// TIA Portal project "FS-DS-09" (V16) (continued)
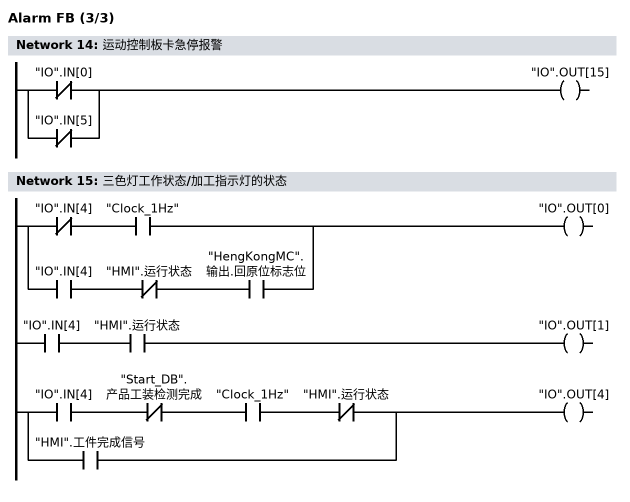
   RUNG wire#powerrail
      I_Contact( "IO".IN[0] )
      wire#w1
      Coil( "IO".OUT[15] )
   END_RUNG
   RUNG wire#powerrail
      I_Contact( "IO".IN[5] )
   END_RUNG wire#w1
   // the same network as SCL:
   "IO".OUT[15] := NOT "IO".IN[0] OR NOT "IO".IN[5];
END_REGION

REGION Network 15: 三色灯工作状态/加工指示灯的状态
   RUNG wire#powerrail
      I_Contact( "IO".IN[4] )
      Contact( "Clock_1Hz" )
      wire#w1
      Coil( "IO".OUT[0] )
   END_RUNG
   RUNG wire#powerrail
      Contact( "IO".IN[4] )
      I_Contact( "HMI".运行状态 )
      Contact( "HengKongMC".输出.回原位标志位 )
   END_RUNG wire#w1
   RUNG wire#powerrail
      Contact( "IO".IN[4] )
      Contact( "HMI".运行状态 )
      Coil( "IO".OUT[1] )
   END_RUNG
   RUNG wire#powerrail
      Contact( "IO".IN[4] )
      I_Contact( "Start_DB".产品工装检测完成 )
      Contact( "Clock_1Hz" )
      I_Contact( "HMI".运行状态 )
      wire#w2
      Coil( "IO".OUT[4] )
   END_RUNG
   RUNG wire#powerrail
      Contact( "HMI".工件完成信号 )
   END_RUNG wire#w2
   // the same network as SCL:
   "IO".OUT[0] := (NOT "IO".IN[4] AND "Clock_1Hz") OR ("IO".IN[4] AND NOT "HMI".运行状态 AND "HengKongMC".输出.回原位标志位);
   "IO".OUT[1] := "IO".IN[4] AND "HMI".运行状态;
   "IO".OUT[4] := ("IO".IN[4] AND NOT "Start_DB".产品工装检测完成 AND "Clock_1Hz" AND NOT "HMI".运行状态) OR "HMI".工件完成信号;
END_REGION
END_FUNCTION_BLOCK

// folder: Control

FUNCTION_BLOCK "Control FB"   // FB2, LAD
{ S7_Optimized_Access := 'TRUE' }
VERSION : 0.1
   VAR
      功能块_Instance : "AM/UM";
      功能块_Instance_1 : "AM/UM";
      功能块_Instance_2 : "AM/UM";
      功能块_Instance_3 : "AM/UM";
      功能块_Instance_4 : "AM/UM";
      功能块_Instance_5 : "AM/UM";
      功能块_Instance_6 : "AM/UM";
      功能块_Instance_7 : "AM/UM";
      IEC_Timer_0_Instance : TON_TIME;
      F_TRIG_Instance : F_TRIG;
      "AM/UM_1_Instance" : "AM/UM_1";
   END_VAR
BEGIN

REGION Network 1: Y1供料器有料输出
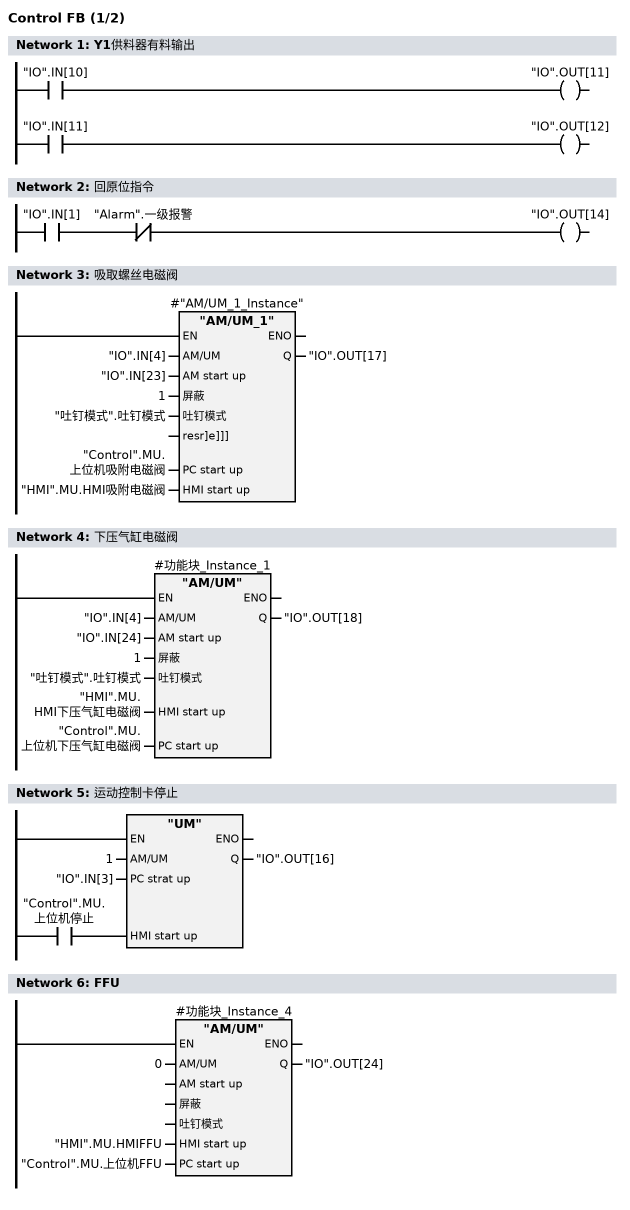
   RUNG wire#powerrail
      Contact( "IO".IN[10] )
      Coil( "IO".OUT[11] )
   END_RUNG
   RUNG wire#powerrail
      Contact( "IO".IN[11] )
      Coil( "IO".OUT[12] )
   END_RUNG
   // the same network as SCL:
   "IO".OUT[11] := "IO".IN[10];
   "IO".OUT[12] := "IO".IN[11];
END_REGION

REGION Network 2: 回原位指令
   RUNG wire#powerrail
      Contact( "IO".IN[1] )
      I_Contact( "Alarm".一级报警 )
      Coil( "IO".OUT[14] )
   END_RUNG
   // the same network as SCL:
   "IO".OUT[14] := "IO".IN[1] AND NOT "Alarm".一级报警;
END_REGION

REGION Network 3: 吸取螺丝电磁阀
   RUNG wire#powerrail
      #"AM/UM_1_Instance"("AM/UM" := "IO".IN[4], "AM start up" := "IO".IN[23], 屏蔽 := 1, 吐钉模式 := "吐钉模式".吐钉模式, "PC start up" := "Control".MU.上位机吸附电磁阀, "HMI start up" := "HMI".MU.HMI吸附电磁阀, Q => "IO".OUT[17], "resr]e]]]" :=)
   END_RUNG
   // the same network as SCL:
   #"AM/UM_1_Instance"("AM/UM" := "IO".IN[4],   // "AM/UM_1"
                       "AM start up" := "IO".IN[23],
                       屏蔽 := 1,
                       吐钉模式 := "吐钉模式".吐钉模式,
                       "PC start up" := "Control".MU.上位机吸附电磁阀,
                       "HMI start up" := "HMI".MU.HMI吸附电磁阀,
                       Q => "IO".OUT[17]);
END_REGION

REGION Network 4: 下压气缸电磁阀
   RUNG wire#powerrail
      #功能块_Instance_1("AM/UM" := "IO".IN[4], "AM start up" := "IO".IN[24], 屏蔽 := 1, 吐钉模式 := "吐钉模式".吐钉模式, "HMI start up" := "HMI".MU.HMI下压气缸电磁阀, "PC start up" := "Control".MU.上位机下压气缸电磁阀, Q => "IO".OUT[18])
   END_RUNG
   // the same network as SCL:
   #功能块_Instance_1("AM/UM" := "IO".IN[4],   // "AM/UM"
                   "AM start up" := "IO".IN[24],
                   屏蔽 := 1,
                   吐钉模式 := "吐钉模式".吐钉模式,
                   "HMI start up" := "HMI".MU.HMI下压气缸电磁阀,
                   "PC start up" := "Control".MU.上位机下压气缸电磁阀,
                   Q => "IO".OUT[18]);
END_REGION

REGION Network 5: 运动控制卡停止
   RUNG wire#powerrail
      "UM"("HMI start up" := wire#w1, "AM/UM" := 1, "PC strat up" := "IO".IN[3], Q => "IO".OUT[16])
   END_RUNG
   RUNG wire#powerrail
      Contact( "Control".MU.上位机停止 )
   END_RUNG wire#w1
   // the same network as SCL:
   "UM"("AM/UM" := 1, "PC strat up" := "IO".IN[3], "HMI start up" := "Control".MU.上位机停止, Q => "IO".OUT[16]);
END_REGION

REGION Network 6: FFU
   RUNG wire#powerrail
      #功能块_Instance_4("AM/UM" := 0, "AM start up" :=, 屏蔽 :=, 吐钉模式 :=, "HMI start up" := "HMI".MU.HMIFFU, "PC start up" := "Control".MU.上位机FFU, Q => "IO".OUT[24])
   END_RUNG
   // the same network as SCL:
   #功能块_Instance_4("AM/UM" := 0,   // "AM/UM"
                   "HMI start up" := "HMI".MU.HMIFFU,
                   "PC start up" := "Control".MU.上位机FFU,
                   Q => "IO".OUT[24]);
END_REGION

REGION Network 7: 照明
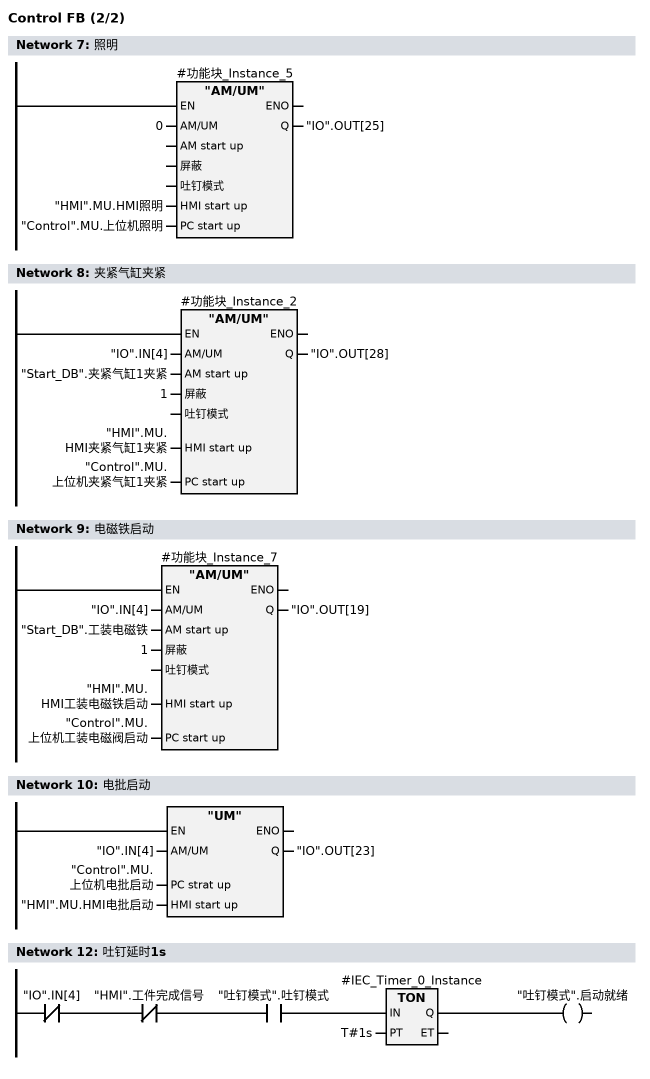
   RUNG wire#powerrail
      #功能块_Instance_5("AM/UM" := 0, "AM start up" :=, 屏蔽 :=, 吐钉模式 :=, "HMI start up" := "HMI".MU.HMI照明, "PC start up" := "Control".MU.上位机照明, Q => "IO".OUT[25])
   END_RUNG
   // the same network as SCL:
   #功能块_Instance_5("AM/UM" := 0,   // "AM/UM"
                   "HMI start up" := "HMI".MU.HMI照明,
                   "PC start up" := "Control".MU.上位机照明,
                   Q => "IO".OUT[25]);
END_REGION

REGION Network 8: 夹紧气缸夹紧
   RUNG wire#powerrail
      #功能块_Instance_2("AM/UM" := "IO".IN[4], "AM start up" := "Start_DB".夹紧气缸1夹紧, 屏蔽 := 1, 吐钉模式 :=, "HMI start up" := "HMI".MU.HMI夹紧气缸1夹紧, "PC start up" := "Control".MU.上位机夹紧气缸1夹紧, Q => "IO".OUT[28])
   END_RUNG
   // the same network as SCL:
   #功能块_Instance_2("AM/UM" := "IO".IN[4],   // "AM/UM"
                   "AM start up" := "Start_DB".夹紧气缸1夹紧,
                   屏蔽 := 1,
                   "HMI start up" := "HMI".MU.HMI夹紧气缸1夹紧,
                   "PC start up" := "Control".MU.上位机夹紧气缸1夹紧,
                   Q => "IO".OUT[28]);
END_REGION

REGION Network 9: 电磁铁启动
   RUNG wire#powerrail
      #功能块_Instance_7("AM/UM" := "IO".IN[4], "AM start up" := "Start_DB".工装电磁铁, 屏蔽 := 1, 吐钉模式 :=, "HMI start up" := "HMI".MU.HMI工装电磁铁启动, "PC start up" := "Control".MU.上位机工装电磁阀启动, Q => "IO".OUT[19])
   END_RUNG
   // the same network as SCL:
   #功能块_Instance_7("AM/UM" := "IO".IN[4],   // "AM/UM"
                   "AM start up" := "Start_DB".工装电磁铁,
                   屏蔽 := 1,
                   "HMI start up" := "HMI".MU.HMI工装电磁铁启动,
                   "PC start up" := "Control".MU.上位机工装电磁阀启动,
                   Q => "IO".OUT[19]);
END_REGION

REGION Network 10: 电批启动
   RUNG wire#powerrail
      "UM"("AM/UM" := "IO".IN[4], "PC strat up" := "Control".MU.上位机电批启动, "HMI start up" := "HMI".MU.HMI电批启动, Q => "IO".OUT[23])
   END_RUNG
   // the same network as SCL:
   "UM"("AM/UM" := "IO".IN[4],
        "PC strat up" := "Control".MU.上位机电批启动,
        "HMI start up" := "HMI".MU.HMI电批启动,
        Q => "IO".OUT[23]);
END_REGION

REGION Network 12: 吐钉延时1s
   #IEC_Timer_0_Instance(IN := NOT "IO".IN[4] AND NOT "HMI".工件完成信号 AND "吐钉模式".吐钉模式, PT := T#1s);   // TON
   "吐钉模式".启动就绪 := #IEC_Timer_0_Instance.Q;
END_REGION

REGION Network 13 (SCL): 完成后 复位
   #F_TRIG_Instance(CLK:="HengKongMC".输出.下压气缸信号,
                    Q=>"吐钉模式".下压气缸复位信号);
   IF "吐钉模式".下压气缸复位信号 OR  "IO".IN[1] THEN
       "吐钉模式".吐钉模式 := 0;
   END_IF;
END_REGION
END_FUNCTION_BLOCK

FUNCTION_BLOCK "Start"   // FB4, LAD
{ S7_Optimized_Access := 'TRUE' }
VERSION : 0.1
   VAR_OUTPUT
      夹紧气缸1夹紧 : Bool;
      夹紧气缸2夹紧 : Bool;
      工装电磁铁 : Bool;
   END_VAR
   VAR
      产品工装检测完成 : Bool;
      气缸夹紧完成 : Bool;
      P1 : Bool;
      P2 : Bool;
      RecipeExport_Instance : RecipeExport;
      RecipeImport_Instance : RecipeImport;
   END_VAR
   VAR_TEMP   // added for the SCL form of the ladder/FBD networks
      _w1 : Bool;
      _w2 : Bool;
   END_VAR
BEGIN

REGION Network 1: 启动1序/停止序
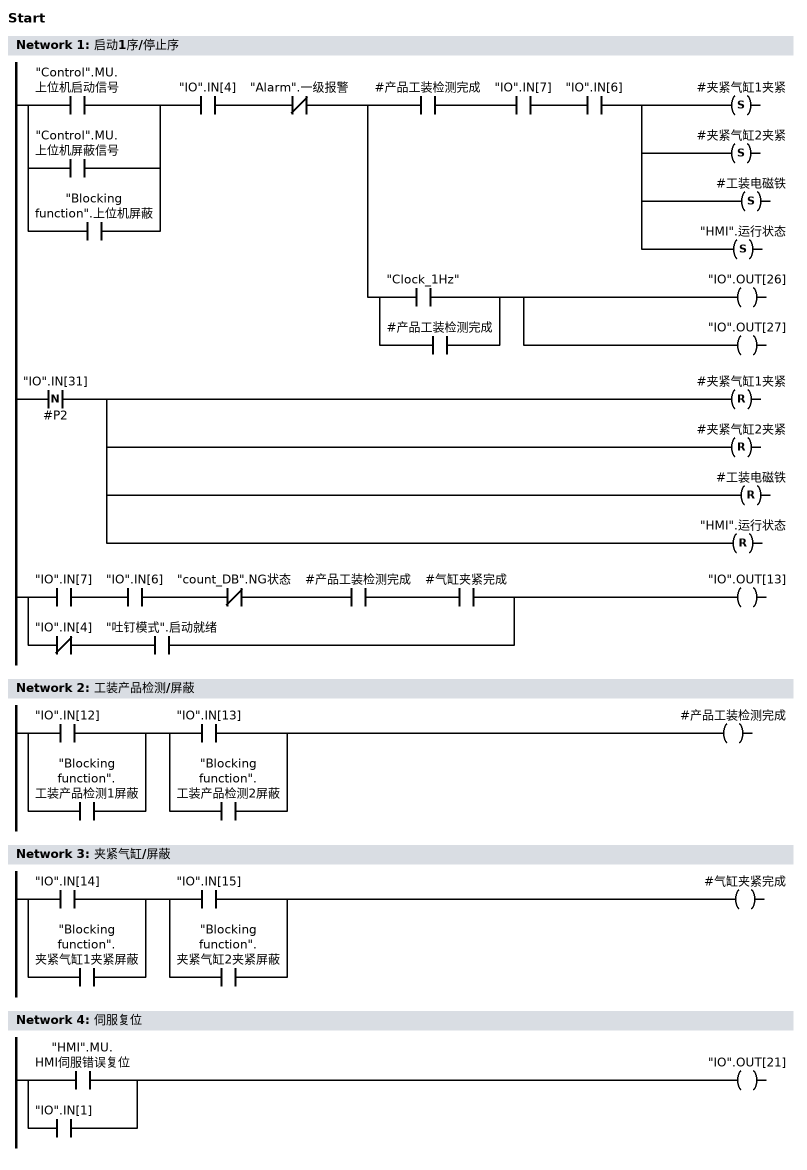
   RUNG wire#powerrail
      Contact( "Control".MU.上位机启动信号 )
      wire#w1
      Contact( "IO".IN[4] )
      I_Contact( "Alarm".一级报警 )
      wire#w2
      Contact( #产品工装检测完成 )
      Contact( "IO".IN[7] )
      Contact( "IO".IN[6] )
      wire#w3
      S_Coil( #夹紧气缸1夹紧 )
   END_RUNG
   RUNG wire#powerrail
      Contact( "Control".MU.上位机屏蔽信号 )
   END_RUNG wire#w1
   RUNG wire#powerrail
      Contact( "Blocking function".上位机屏蔽 )
   END_RUNG wire#w1
   RUNG wire#w3
      S_Coil( #夹紧气缸2夹紧 )
   END_RUNG
   RUNG wire#w3
      S_Coil( #工装电磁铁 )
   END_RUNG
   RUNG wire#w3
      S_Coil( "HMI".运行状态 )
   END_RUNG
   RUNG wire#w2
      Contact( "Clock_1Hz" )
      wire#w4
      Coil( "IO".OUT[26] )
   END_RUNG
   RUNG wire#w2
      Contact( #产品工装检测完成 )
   END_RUNG wire#w4
   RUNG wire#w4
      Coil( "IO".OUT[27] )
   END_RUNG
   RUNG wire#powerrail
      N_Contact(operand := "IO".IN[31], bit := #P2)
      wire#w5
      R_Coil( #夹紧气缸1夹紧 )
   END_RUNG
   RUNG wire#w5
      R_Coil( #夹紧气缸2夹紧 )
   END_RUNG
   RUNG wire#w5
      R_Coil( #工装电磁铁 )
   END_RUNG
   RUNG wire#w5
      R_Coil( "HMI".运行状态 )
   END_RUNG
   RUNG wire#powerrail
      Contact( "IO".IN[7] )
      Contact( "IO".IN[6] )
      I_Contact( "count_DB".NG状态 )
      Contact( #产品工装检测完成 )
      Contact( #气缸夹紧完成 )
      wire#w6
      Coil( "IO".OUT[13] )
   END_RUNG
   RUNG wire#powerrail
      I_Contact( "IO".IN[4] )
      Contact( "吐钉模式".启动就绪 )
   END_RUNG wire#w6
   // the same network as SCL:
   #_w1 := ("Control".MU.上位机启动信号 OR "Control".MU.上位机屏蔽信号 OR "Blocking function".上位机屏蔽) AND "IO".IN[4] AND NOT "Alarm".一级报警;
   IF #_w1 AND #产品工装检测完成 AND "IO".IN[7] AND "IO".IN[6] THEN
       #夹紧气缸1夹紧 := TRUE;
       #夹紧气缸2夹紧 := TRUE;
       #工装电磁铁 := TRUE;
       "HMI".运行状态 := TRUE;
   END_IF;
   "IO".OUT[26] := #_w1 AND ("Clock_1Hz" OR #产品工装检测完成);
   "IO".OUT[27] := #_w1 AND ("Clock_1Hz" OR #产品工装检测完成);
   #_w2 := NOT "IO".IN[31] AND #P2;   // falling edge of "IO".IN[31]
   #P2 := "IO".IN[31];
   IF #_w2 THEN
       #夹紧气缸1夹紧 := FALSE;
       #夹紧气缸2夹紧 := FALSE;
       #工装电磁铁 := FALSE;
       "HMI".运行状态 := FALSE;
   END_IF;
   "IO".OUT[13] := ("IO".IN[7] AND "IO".IN[6] AND NOT "count_DB".NG状态 AND #产品工装检测完成 AND #气缸夹紧完成) OR (NOT "IO".IN[4] AND "吐钉模式".启动就绪);
END_REGION

REGION Network 2: 工装产品检测/屏蔽
   RUNG wire#powerrail
      Contact( "IO".IN[12] )
      wire#w1
      Contact( "IO".IN[13] )
      wire#w2
      Coil( #产品工装检测完成 )
   END_RUNG
   RUNG wire#powerrail
      Contact( "Blocking function".工装产品检测1屏蔽 )
   END_RUNG wire#w1
   RUNG wire#w1
      Contact( "Blocking function".工装产品检测2屏蔽 )
   END_RUNG wire#w2
   // the same network as SCL:
   #产品工装检测完成 := ("IO".IN[12] OR "Blocking function".工装产品检测1屏蔽) AND ("IO".IN[13] OR "Blocking function".工装产品检测2屏蔽);
END_REGION

REGION Network 3: 夹紧气缸/屏蔽
   RUNG wire#powerrail
      Contact( "IO".IN[14] )
      wire#w1
      Contact( "IO".IN[15] )
      wire#w2
      Coil( #气缸夹紧完成 )
   END_RUNG
   RUNG wire#powerrail
      Contact( "Blocking function".夹紧气缸1夹紧屏蔽 )
   END_RUNG wire#w1
   RUNG wire#w1
      Contact( "Blocking function".夹紧气缸2夹紧屏蔽 )
   END_RUNG wire#w2
   // the same network as SCL:
   #气缸夹紧完成 := ("IO".IN[14] OR "Blocking function".夹紧气缸1夹紧屏蔽) AND ("IO".IN[15] OR "Blocking function".夹紧气缸2夹紧屏蔽);
END_REGION

REGION Network 4: 伺服复位
   RUNG wire#powerrail
      Contact( "HMI".MU.HMI伺服错误复位 )
      wire#w1
      Coil( "IO".OUT[21] )
   END_RUNG
   RUNG wire#powerrail
      Contact( "IO".IN[1] )
   END_RUNG wire#w1
   // the same network as SCL:
   "IO".OUT[21] := "HMI".MU.HMI伺服错误复位 OR "IO".IN[1];
END_REGION
END_FUNCTION_BLOCK

FUNCTION_BLOCK "AM/UM"   // FB5, LAD
{ S7_Optimized_Access := 'TRUE' }
VERSION : 0.1
   VAR_INPUT
      "AM/UM" : Bool;   // 手动自动
      "AM start up" : Bool;   // 自动启动
      屏蔽 : Bool;   // 屏蔽0
      吐钉模式 : Bool;
   END_VAR
   VAR_OUTPUT
      Q : Bool;   // 功能输出
   END_VAR
   VAR_IN_OUT
      "HMI start up" : Bool;   // HMI启动
      "PC start up" : Bool;   // 上位机启动
   END_VAR
   VAR
      F_TRIG_Instance : F_TRIG;
   END_VAR
BEGIN

REGION Network 1: 功能输出
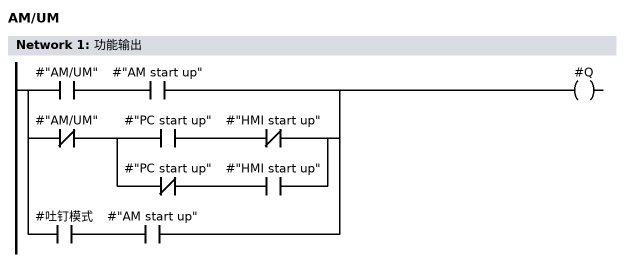
   RUNG wire#powerrail
      Contact( #"AM/UM" )
      Contact( #"AM start up" )
      wire#w1
      Coil( #Q )
   END_RUNG
   RUNG wire#powerrail
      I_Contact( #"AM/UM" )
      wire#w2
      Contact( #"PC start up" )
      I_Contact( #"HMI start up" )
   END_RUNG wire#w1
   RUNG wire#w2
      I_Contact( #"PC start up" )
      Contact( #"HMI start up" )
   END_RUNG wire#w1
   RUNG wire#powerrail
      Contact( #吐钉模式 )
      Contact( #"AM start up" )
   END_RUNG wire#w1
   // the same network as SCL:
   #Q := (#"AM/UM" AND #"AM start up") OR (NOT #"AM/UM" AND ((#"PC start up" AND NOT #"HMI start up") OR (NOT #"PC start up" AND #"HMI start up"))) OR (#吐钉模式 AND #"AM start up");
END_REGION

REGION Network 2 (SCL): HMI启动
   IF #屏蔽 THEN
       IF #"AM/UM" = 1 THEN
           #"HMI start up" := 0;
           #"PC start up":=0
           ;
       END_IF;
   END_IF;
END_REGION
END_FUNCTION_BLOCK

FUNCTION_BLOCK "count"   // FB7, LAD
{ S7_Optimized_Access := 'TRUE' }
VERSION : 0.1
// 计数OK/NG/累计/ 合格率
   VAR_INPUT
      CE : Bool;   // 清零
      "AM/UM" : Bool;   // 手动自动
   END_VAR
   VAR_OUTPUT
      "OK Screw mumber" : Int;   // 拧到第几个螺丝
      "OK screw" : Bool;   // 工件加工合格
      "NG screw" : Bool;   // 工件加工不合格
      OK_1 : Real;
      NG_1 : Real;
      "NG Screw mumber_1" : Int;   // 拧到第几个螺丝
   END_VAR
   VAR_IN_OUT
      OK : Bool;   // 电批合格信号
      "OK+NG" : Real;
      "OK/NG%" : Real;
      NG : Bool;   // 电批不合格信号
      Number : Int;   // 数量（锁螺丝数量）
   END_VAR
   VAR RETAIN
      IEC_Counter_0_Instance : CTU_INT;
      IEC_Counter_0_Instance_1 : CTU_INT;
      P1 : Bool;
      P2 : Bool;
   END_VAR
   VAR
      P3 : Bool;
      P4 : Bool;
      P5 : Bool;
      P6 : Bool;
      P7 : Bool;
      p8 : Bool;
      P9 : Bool;
      P10 : Bool;
      P11 : Bool;
      P12 : Bool;
      P13 : Bool;
      螺丝加工完成 : Bool;
   END_VAR
   VAR RETAIN
      IEC_Counter_0_Instance_2 : CTU_INT;
   END_VAR
   VAR
      "NG Screw mumber" : Int;   // 拧到第几个螺丝
      加工状态对比 : Word := 16#F1;
      NG状态 : Bool;
      重打 : Bool;
   END_VAR
   VAR_TEMP   // added for the SCL form of the ladder/FBD networks
      _w1 : Bool;
      _w2 : Bool;
      _w3 : Bool;
      _w4 : Bool;
      _w5 : Bool;
      _w6 : Bool;
      _w7 : Bool;
   END_VAR
BEGIN

REGION Network 1 (SCL)
   // 产品计数和合格率
   #"OK+NG" :=  #OK_1 + #NG_1;//累计
   #"OK/NG%" := (#OK_1 / #"OK+NG"*100);//合格率
   //IF #"OK+NG" = 32760 OR #CE THEN
      // #IEC_Counter_0_Instance.R := 1;
      // #IEC_Counter_0_Instance_1.R := 1;
   //END_IF;//清零
   IF #NG THEN
       #"NG Screw mumber_1" := #"OK Screw mumber" + #"NG Screw mumber";
   ELSE
       #"NG Screw mumber_1" := 0;
   END_IF;
END_REGION

REGION Network 2: 合格计数
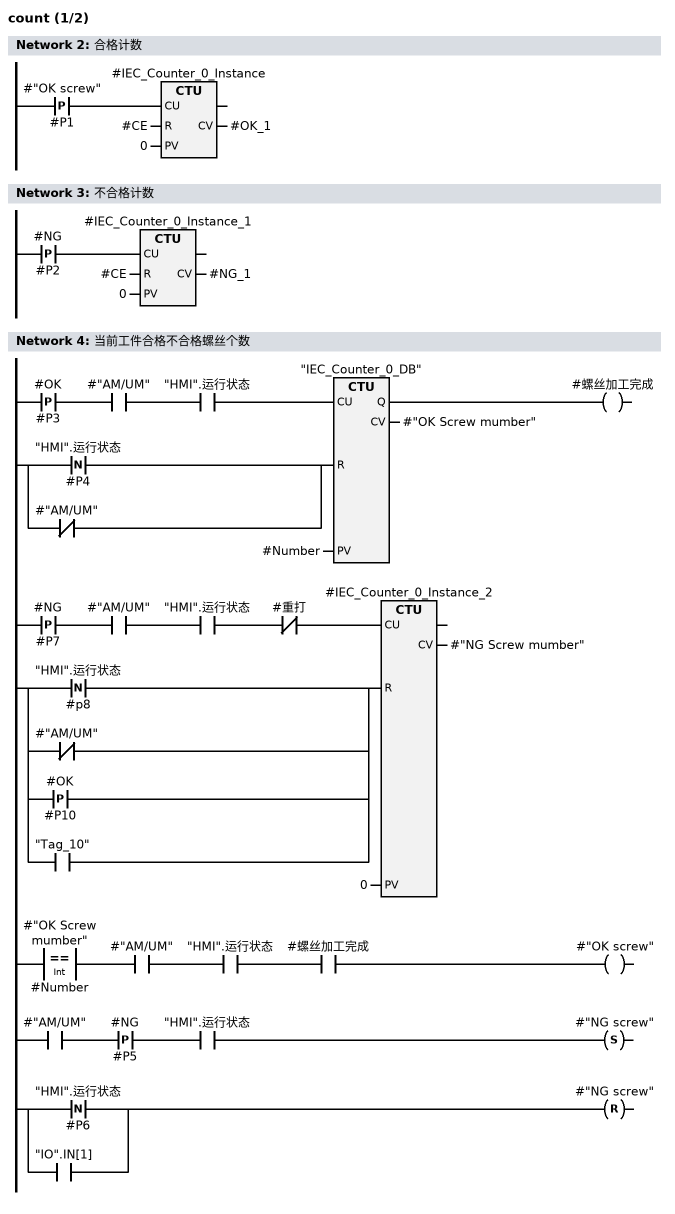
   #_w1 := #"OK screw" AND NOT #P1;   // rising edge of #"OK screw"
   #P1 := #"OK screw";
   #IEC_Counter_0_Instance(CU := #_w1, R := #CE, PV := 0, CV => #OK_1);   // CTU
END_REGION

REGION Network 3: 不合格计数
   #_w1 := #NG AND NOT #P2;   // rising edge of #NG
   #P2 := #NG;
   #IEC_Counter_0_Instance_1(CU := #_w1, R := #CE, PV := 0, CV => #NG_1);   // CTU
END_REGION

REGION Network 4: 当前工件合格不合格螺丝个数
   #_w1 := #OK AND NOT #P3;   // rising edge of #OK
   #P3 := #OK;
   #_w2 := NOT "HMI".运行状态 AND #P4;   // falling edge of "HMI".运行状态
   #P4 := "HMI".运行状态;
   "IEC_Counter_0_DB".CTU(CU := #_w1 AND #"AM/UM" AND "HMI".运行状态,
                          R := #_w2 OR NOT #"AM/UM",
                          PV := #Number,
                          CV => #"OK Screw mumber");
   #螺丝加工完成 := "IEC_Counter_0_DB".Q;
   #_w3 := #NG AND NOT #P7;   // rising edge of #NG
   #P7 := #NG;
   #_w4 := NOT "HMI".运行状态 AND #p8;   // falling edge of "HMI".运行状态
   #p8 := "HMI".运行状态;
   #_w5 := #OK AND NOT #P10;   // rising edge of #OK
   #P10 := #OK;
   #IEC_Counter_0_Instance_2(CU := #_w3 AND #"AM/UM" AND "HMI".运行状态 AND NOT #重打,   // CTU
                           R := #_w4 OR NOT #"AM/UM" OR #_w5 OR "Tag_10",
                           PV := 0,
                           CV => #"NG Screw mumber");
   #"OK screw" := (#"OK Screw mumber" = #Number) AND #"AM/UM" AND "HMI".运行状态 AND #螺丝加工完成;
   #_w6 := #"AM/UM" AND #NG AND NOT #P5;   // rising edge of #NG
   #P5 := #NG;
   IF #_w6 AND "HMI".运行状态 THEN #"NG screw" := TRUE; END_IF;
   #_w7 := NOT "HMI".运行状态 AND #P6;   // falling edge of "HMI".运行状态
   #P6 := "HMI".运行状态;
   IF #_w7 OR "IO".IN[1] THEN #"NG screw" := FALSE; END_IF;
END_REGION

REGION Network 5: 螺丝拧紧NG的状态下重打执行/按面板启动键执行
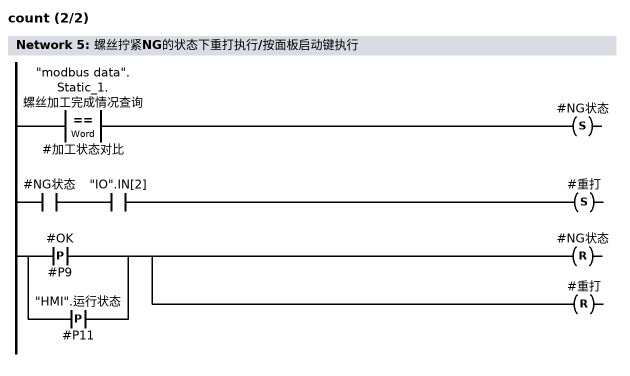
   RUNG wire#powerrail
      { S7_Templates := "SrcType := Word" } EQ_Contact(in1 := "modbus data".Static_1.螺丝加工完成情况查询, in2 := #加工状态对比)
      S_Coil( #NG状态 )
   END_RUNG
   RUNG wire#powerrail
      Contact( #NG状态 )
      Contact( "IO".IN[2] )
      S_Coil( #重打 )
   END_RUNG
   RUNG wire#powerrail
      P_Contact(operand := #OK, bit := #P9)
      wire#w1
      R_Coil( #NG状态 )
   END_RUNG
   RUNG wire#powerrail
      P_Contact(operand := "HMI".运行状态, bit := #P11)
   END_RUNG wire#w1
   RUNG wire#w1
      R_Coil( #重打 )
   END_RUNG
   // the same network as SCL:
   IF "modbus data".Static_1.螺丝加工完成情况查询 = #加工状态对比 THEN #NG状态 := TRUE; END_IF;
   IF #NG状态 AND "IO".IN[2] THEN #重打 := TRUE; END_IF;
   #_w1 := #OK AND NOT #P9;   // rising edge of #OK
   #P9 := #OK;
   #_w2 := "HMI".运行状态 AND NOT #P11;   // rising edge of "HMI".运行状态
   #P11 := "HMI".运行状态;
   IF #_w1 OR #_w2 THEN
       #NG状态 := FALSE;
       #重打 := FALSE;
   END_IF;
END_REGION
END_FUNCTION_BLOCK

FUNCTION_BLOCK "AM/UM_1"   // FB8, LAD
{ S7_Optimized_Access := 'TRUE' }
VERSION : 0.1
   VAR_INPUT
      "AM/UM" : Bool;   // 手动自动
      "AM start up" : Bool;   // 自动启动
      屏蔽 : Bool;   // 屏蔽0
      吐钉模式 : Bool;
      "resr]e]]]" : Bool;
   END_VAR
   VAR_OUTPUT
      Q : Bool;   // 功能输出
   END_VAR
   VAR_IN_OUT
      "PC start up" : Bool;   // 上位机启动
      "HMI start up" : Bool;   // HMI启动
   END_VAR
   VAR
      F_TRIG_Instance : F_TRIG;
      P1 : Bool;
      P2 : Bool;
      P3 : Bool;
      P4 : Bool;
      P5 : Bool;
   END_VAR
   VAR_TEMP   // added for the SCL form of the ladder/FBD networks
      _w1 : Bool;
      _w2 : Bool;
      _w3 : Bool;
   END_VAR
BEGIN

REGION Network 1: 功能输出
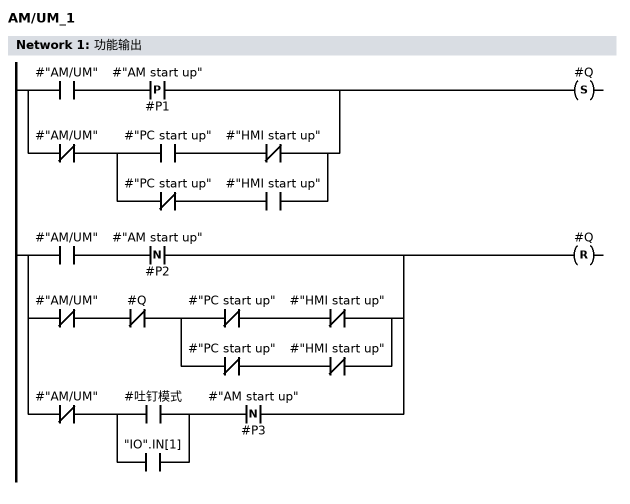
   RUNG wire#powerrail
      Contact( #"AM/UM" )
      P_Contact(operand := #"AM start up", bit := #P1)
      wire#w1
      S_Coil( #Q )
   END_RUNG
   RUNG wire#powerrail
      I_Contact( #"AM/UM" )
      wire#w2
      Contact( #"PC start up" )
      I_Contact( #"HMI start up" )
   END_RUNG wire#w1
   RUNG wire#w2
      I_Contact( #"PC start up" )
      Contact( #"HMI start up" )
   END_RUNG wire#w1
   RUNG wire#powerrail
      Contact( #"AM/UM" )
      N_Contact(operand := #"AM start up", bit := #P2)
      wire#w3
      R_Coil( #Q )
   END_RUNG
   RUNG wire#powerrail
      I_Contact( #"AM/UM" )
      I_Contact( #Q )
      wire#w4
      I_Contact( #"PC start up" )
      I_Contact( #"HMI start up" )
   END_RUNG wire#w3
   RUNG wire#w4
      I_Contact( #"PC start up" )
      I_Contact( #"HMI start up" )
   END_RUNG wire#w3
   RUNG wire#powerrail
      I_Contact( #"AM/UM" )
      wire#w5
      Contact( #吐钉模式 )
      wire#w6
      N_Contact(operand := #"AM start up", bit := #P3)
   END_RUNG wire#w3
   RUNG wire#w5
      Contact( "IO".IN[1] )
   END_RUNG wire#w6
   // the same network as SCL:
   #_w1 := #"AM/UM" AND #"AM start up" AND NOT #P1;   // rising edge of #"AM start up"
   #P1 := #"AM start up";
   IF #_w1 OR (NOT #"AM/UM" AND ((#"PC start up" AND NOT #"HMI start up") OR (NOT #"PC start up" AND #"HMI start up"))) THEN
       #Q := TRUE;
   END_IF;
   #_w2 := #"AM/UM" AND NOT #"AM start up" AND #P2;   // falling edge of #"AM start up"
   #P2 := #"AM start up";
   #_w3 := NOT #"AM/UM" AND (#吐钉模式 OR "IO".IN[1]) AND NOT #"AM start up" AND #P3;   // falling edge of #"AM start up"
   #P3 := #"AM start up";
   IF #_w2 OR (NOT #"AM/UM" AND NOT #Q AND ((NOT #"PC start up" AND NOT #"HMI start up") OR (NOT #"PC start up" AND NOT #"HMI start up"))) OR #_w3 THEN
       #Q := FALSE;
   END_IF;
END_REGION

REGION Network 2 (SCL): HMI启动
   IF #屏蔽 THEN
       IF #"AM/UM" = 1 THEN
           #"HMI start up" := 0;
           #"PC start up" := 0;
       END_IF;
   END_IF;
END_REGION
END_FUNCTION_BLOCK

FUNCTION "UM" : Void   // FC2, LAD
{ S7_Optimized_Access := 'TRUE' }
VERSION : 0.1
   VAR_INPUT
      "AM/UM" : Bool;
      "PC strat up" : Bool;
      "HMI start up" : Bool;
   END_VAR
   VAR_OUTPUT
      Q : Bool;
   END_VAR
BEGIN

REGION Network 1
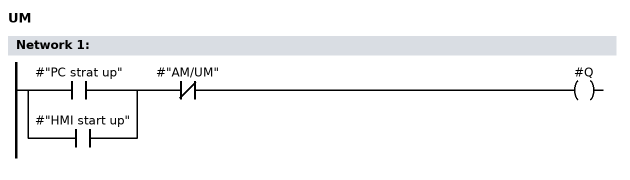
   RUNG wire#powerrail
      Contact( #"PC strat up" )
      wire#w1
      I_Contact( #"AM/UM" )
      Coil( #Q )
   END_RUNG
   RUNG wire#powerrail
      Contact( #"HMI start up" )
   END_RUNG wire#w1
   // the same network as SCL:
   #Q := (#"PC strat up" OR #"HMI start up") AND NOT #"AM/UM";
END_REGION
END_FUNCTION

// folder: DATA

FUNCTION "Data" : Void   // FC1, SCL
{ S7_Optimized_Access := 'TRUE' }
VERSION : 0.1
BEGIN
   REGION IN
       "IO".IN[0] := "操作面板急停";
       "IO".IN[1] := "回原位";
       "IO".IN[2] := "启动按钮";
       "IO".IN[3] := "停止按钮";
       "IO".IN[4] := "手动/自动";
       "IO".IN[5] := "按钮盒急停";
       "IO".IN[6] := "左启动";
       "IO".IN[7] := "右启动";
       "IO".IN[8] := "备用";
       "IO".IN[9] := "光幕";
       "IO".IN[10] := "Y1供料器有料";
       "IO".IN[11] := "Y2供料器有料";
       "IO".IN[12] := "1#工装产品信号";
       "IO".IN[13] := "2#工装产品信号";
       "IO".IN[14] := "气夹气缸到位2";
       "IO".IN[15] := "气夹气缸到位1";
       "IO".IN[16] := "工具错误";
       "IO".IN[17] := "工具拧紧OK";
       "IO".IN[18] := "工具拧紧NG";
       "IO".IN[19] := "工具准备好";
       "IO".IN[20] := "工具运行";
       "IO".IN[21] := "气源压力检测";
       "IO".IN[22] := "光栅屏蔽对射开关";
       "IO".IN[23] := "吸附信号";
       "IO".IN[24] := "电批下压气缸下压信号";
       "IO".IN[25] := "安全门";
       "IO".IN[26] := "回原位中";
       "IO".IN[27] := "回原位完成";
       "IO".IN[28] := "X轴故障报警";
       "IO".IN[29] := "Y轴故障报警";
       "IO".IN[30] := "Z轴故障报警";
       "IO".IN[31] := "运动控制卡完成/释放夹紧气缸";
       "IO".IN[32] := "备用_3";
       "IO".IN[33] := "备用_4";
       "IO".IN[34] := "备用_5";
       "IO".IN[35] := "备用_6";
       "IO".IN[36] := "备用_7";
       "IO".IN[37] := "备用_8";
       "IO".IN[38] := 0;
       "IO".IN[39] := 0;
       "IO".IN[40] := 0;

   END_REGION
   REGION OUT
       "三色灯黄色" := "IO".OUT[0];
       "IO".OUT[1] := "三色灯绿色" := "IO".OUT[1];
       "三色灯红色" := "IO".OUT[2];
       "三色灯蜂鸣器" := "IO".OUT[3];
       "绿色半球指示灯" := "IO".OUT[4];
       "红色半球指示灯" := "IO".OUT[5];
       "运动控制卡任务选择1" := "IO".OUT[6];
       "运动控制卡任务选择2" := "IO".OUT[7];
       "运动控制卡任务选择3" := "IO".OUT[8];
       "运动控制卡任务选择4" := "IO".OUT[9];
       "运动控制卡任务选择5" := "IO".OUT[10];
       "Y1供料器有料输出" := "IO".OUT[11];
       "Y2供料器有料输出" := "IO".OUT[12];
       "运动控制卡启动" := "IO".OUT[13];
       "运动控制卡复位" := "IO".OUT[14];
       "运动控制卡紧急停止" := "IO".OUT[15];
       "运动控制卡停止" := "IO".OUT[16];
       "吸取螺丝电磁阀" := "IO".OUT[17];
       "下压气缸电磁阀" := "IO".OUT[18];
       "工装电磁铁" := "IO".OUT[19];
       "光栅报警" := "IO".OUT[20];
       "伺服复位" := "IO".OUT[21];
       "电批急停" := "IO".OUT[22];
       "电批测试启动" := "IO".OUT[23];
       "FFU" := "IO".OUT[24];
       "照明" := "IO".OUT[25];
       "左启动指示灯" := "IO".OUT[26];
       "右启动指示灯" := "IO".OUT[27];
       "夹紧气缸夹紧" := "IO".OUT[28];
       "伺服报警" := "IO".OUT[29];
       "备用_5(1)" := "IO".OUT[30];
       "备用_6(1)" := "IO".OUT[31];
       "备用_7(1)" := "IO".OUT[32];
       "备用_8(1)" := "IO".OUT[33];
       "IO".OUT[34] := 0;
       "IO".OUT[35] := 0;
       "IO".OUT[36] := 0;
       "IO".OUT[37] := 0;
       "IO".OUT[38] := 0;
       "IO".OUT[39] := 0;
       "IO".OUT[40] := 0;

   END_REGION
END_FUNCTION

// folder: Mudbus TCP

FUNCTION_BLOCK "modbus tcp"   // FB1, LAD
{ S7_Optimized_Access := 'TRUE' }
VERSION : 0.1
   VAR
      "DONE 11" : Bool;
      "BUSY 11" : Bool;
      ERROR11 : Bool;
      "DONE 12" : Bool;
      "BUSY 12" : Bool;
      ERROR12 : Bool;
      "DONE 13" : Bool;
      "BUSY 13" : Bool;
      ERROR13 : Bool;
      "DONE 14" : Bool;
      "BUSY 14" : Bool;
      ERROR14 : Bool;
      "DONE 15" : Bool;
      "BUSY 15" : Bool;
      ERROR15 : Bool;
      "DONE 16" : Bool;
      "BUSY 16" : Bool;
      ERROR16 : Bool;
      "DONE 17" : Bool;
      "BUSY 17" : Bool;
      ERROR17 : Bool;
      "DONE 18" : Bool;
      "BUSY 18" : Bool;
      ERROR18 : Bool;
      "DONE 19" : Bool;
      "BUSY 19" : Bool;
      ERROR19 : Bool;
      CF1 : Bool;
      CF2 : Bool;
      CF3 : Bool;
      CF4 : Bool;
      CF5 : Bool;
      CF6 : Bool;
      CF7 : Bool;
      CF8 : Bool;
      CF9 : Bool;
      IEC_Timer_0_Instance_2 : TP_TIME;
      P1 : Bool;
      P2 : Bool;
      P3 : Bool;
      p4 : Bool;
      p5 : Bool;
      p6 : Bool;
      p7 : Bool;
      IEC_Timer_0_Instance : TP_TIME;
      回原位标志位写入 : Bool;
      "1" : Bool := 1;
      "0" : Bool := 0;
      IEC_Timer_0_Instance_1 : TON_TIME;
   END_VAR
   VAR_TEMP   // added for the SCL form of the ladder/FBD networks
      _w1 : Bool;
      _w2 : Bool;
      _w3 : Bool;
      _w4 : Bool;
      _w5 : Bool;
      _w6 : Bool;
   END_VAR
BEGIN

REGION Network 1: 输入
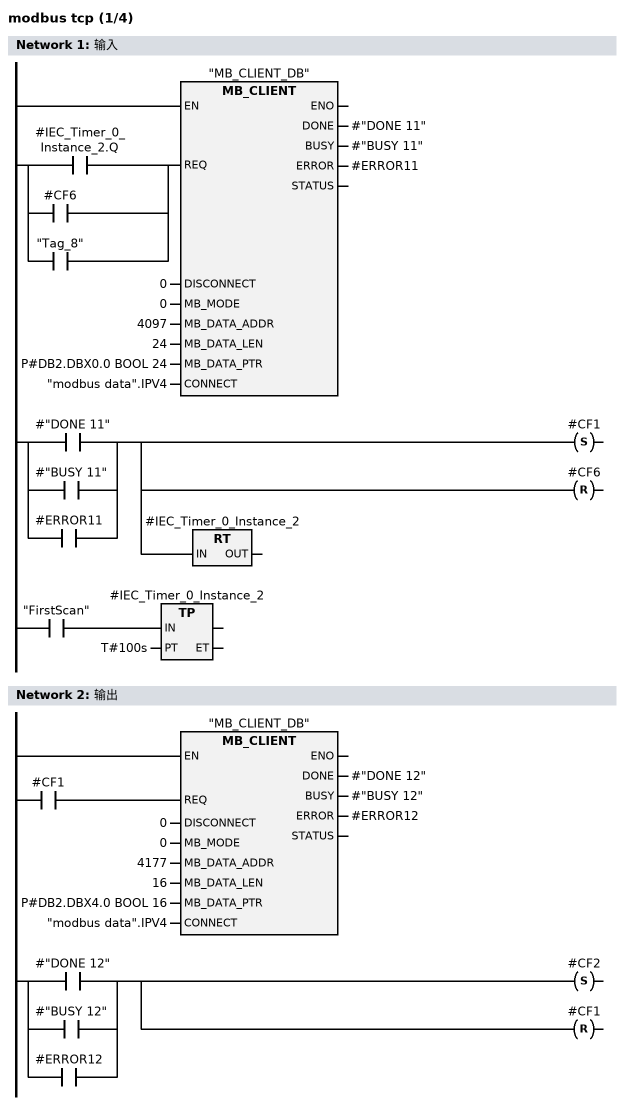
   "MB_CLIENT_DB"(REQ := #IEC_Timer_0_Instance_2.Q OR #CF6 OR "Tag_8",   // MB_CLIENT
                  DISCONNECT := 0,
                  MB_MODE := 0,
                  MB_DATA_ADDR := 4097,
                  MB_DATA_LEN := 24,
                  MB_DATA_PTR := P#DB2.DBX0.0 BOOL 24,
                  CONNECT := "modbus data".IPV4,
                  DONE => #"DONE 11",
                  BUSY => #"BUSY 11",
                  ERROR => #ERROR11);
   #_w1 := #"DONE 11" OR #"BUSY 11" OR #ERROR11;
   IF #_w1 THEN
       #CF1 := TRUE;
       #CF6 := FALSE;
       RESET_TIMER(#IEC_Timer_0_Instance_2);
   END_IF;
   #IEC_Timer_0_Instance_2(IN := "FirstScan", PT := T#100s);   // TP
END_REGION

REGION Network 2: 输出
   "MB_CLIENT_DB"(REQ := #CF1,   // MB_CLIENT
                  DISCONNECT := 0,
                  MB_MODE := 0,
                  MB_DATA_ADDR := 4177,
                  MB_DATA_LEN := 16,
                  MB_DATA_PTR := P#DB2.DBX4.0 BOOL 16,
                  CONNECT := "modbus data".IPV4,
                  DONE => #"DONE 12",
                  BUSY => #"BUSY 12",
                  ERROR => #ERROR12);
   IF #"DONE 12" OR #"BUSY 12" OR #ERROR12 THEN
       #CF2 := TRUE;
       #CF1 := FALSE;
   END_IF;
END_REGION

REGION Network 3: 坐标
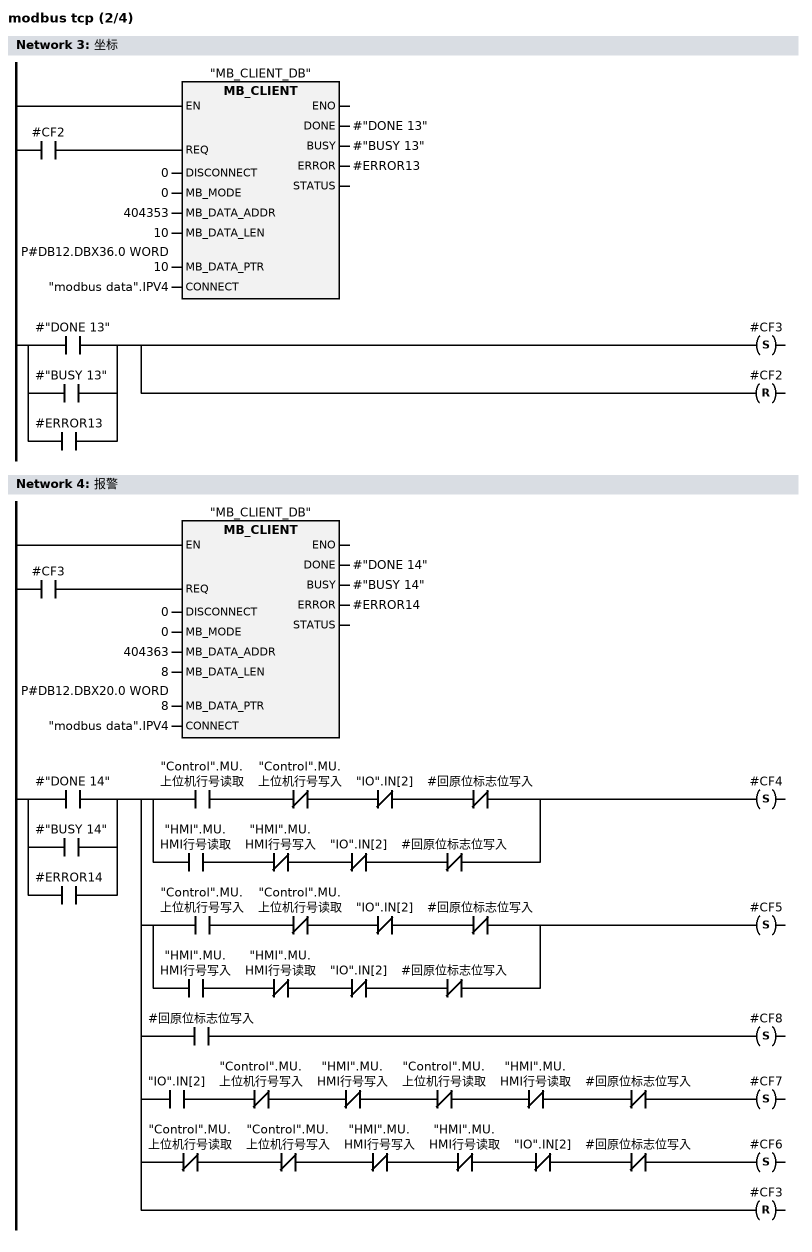
   "MB_CLIENT_DB"(REQ := #CF2,   // MB_CLIENT
                  DISCONNECT := 0,
                  MB_MODE := 0,
                  MB_DATA_ADDR := 404353,
                  MB_DATA_LEN := 10,
                  MB_DATA_PTR := P#DB12.DBX36.0 WORD 10,
                  CONNECT := "modbus data".IPV4,
                  DONE => #"DONE 13",
                  BUSY => #"BUSY 13",
                  ERROR => #ERROR13);
   IF #"DONE 13" OR #"BUSY 13" OR #ERROR13 THEN
       #CF3 := TRUE;
       #CF2 := FALSE;
   END_IF;
END_REGION

REGION Network 4: 报警
   "MB_CLIENT_DB"(REQ := #CF3,   // MB_CLIENT
                  DISCONNECT := 0,
                  MB_MODE := 0,
                  MB_DATA_ADDR := 404363,
                  MB_DATA_LEN := 8,
                  MB_DATA_PTR := P#DB12.DBX20.0 WORD 8,
                  CONNECT := "modbus data".IPV4,
                  DONE => #"DONE 14",
                  BUSY => #"BUSY 14",
                  ERROR => #ERROR14);
   #_w1 := #"DONE 14" OR #"BUSY 14" OR #ERROR14;
   IF #_w1 AND (("Control".MU.上位机行号读取 AND NOT "Control".MU.上位机行号写入 AND NOT "IO".IN[2] AND NOT #回原位标志位写入) OR ("HMI".MU.HMI行号读取 AND NOT "HMI".MU.HMI行号写入 AND NOT "IO".IN[2] AND NOT #回原位标志位写入)) THEN
       #CF4 := TRUE;
   END_IF;
   IF #_w1 AND (("Control".MU.上位机行号写入 AND NOT "Control".MU.上位机行号读取 AND NOT "IO".IN[2] AND NOT #回原位标志位写入) OR ("HMI".MU.HMI行号写入 AND NOT "HMI".MU.HMI行号读取 AND NOT "IO".IN[2] AND NOT #回原位标志位写入)) THEN
       #CF5 := TRUE;
   END_IF;
   IF #_w1 AND #回原位标志位写入 THEN #CF8 := TRUE; END_IF;
   IF #_w1 AND "IO".IN[2] AND NOT "Control".MU.上位机行号写入 AND NOT "HMI".MU.HMI行号写入 AND NOT "Control".MU.上位机行号读取 AND NOT "HMI".MU.HMI行号读取 AND NOT #回原位标志位写入 THEN
       #CF7 := TRUE;
   END_IF;
   IF #_w1 AND NOT "Control".MU.上位机行号读取 AND NOT "Control".MU.上位机行号写入 AND NOT "HMI".MU.HMI行号写入 AND NOT "HMI".MU.HMI行号读取 AND NOT "IO".IN[2] AND NOT #回原位标志位写入 THEN
       #CF6 := TRUE;
   END_IF;
   IF #_w1 THEN #CF3 := FALSE; END_IF;
END_REGION

REGION Network 5: 补螺丝功能读取